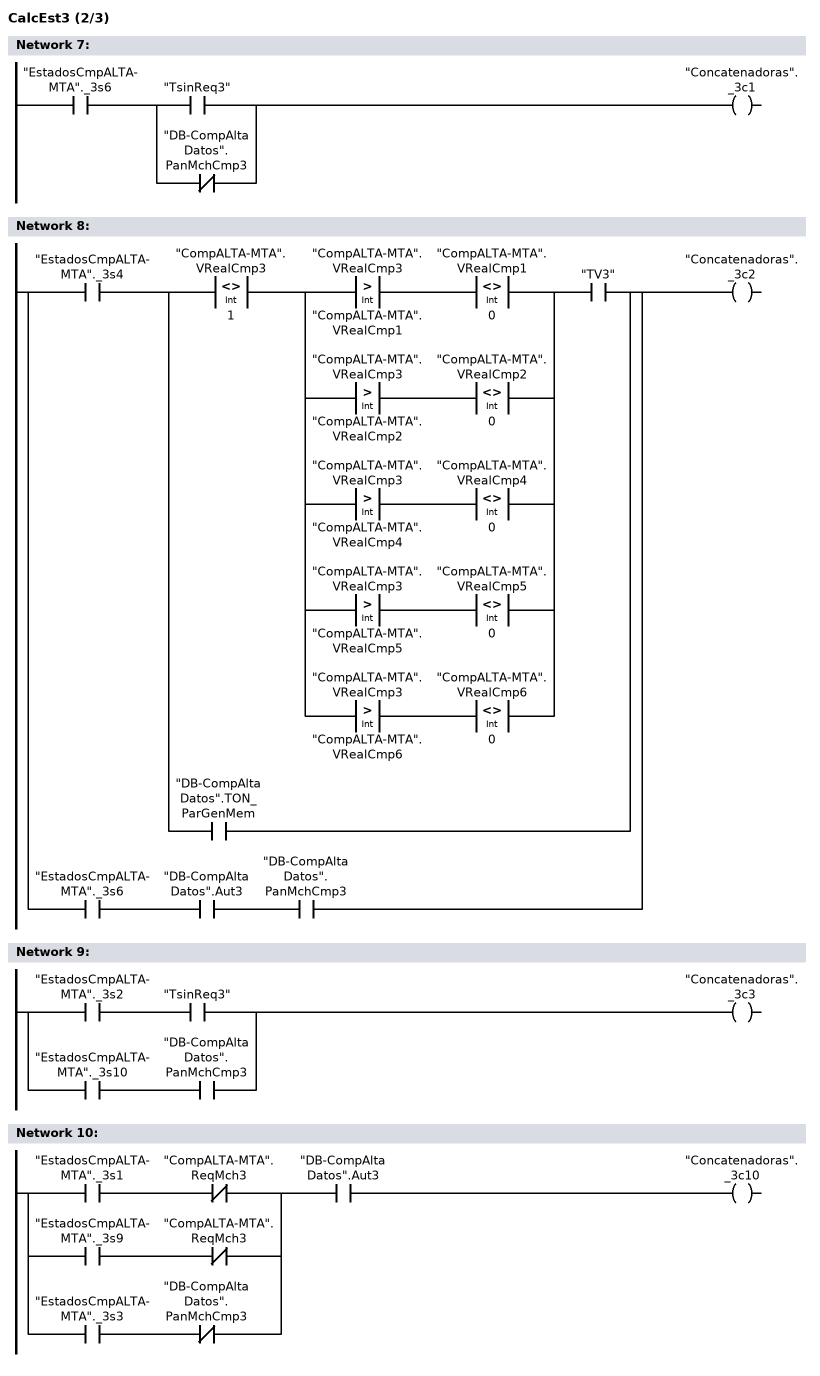
   RUNG wire#powerrail
      Contact( "EstadosCmpALTA-MTA"._3s6 )
      wire#w1
      Contact( "TsinReq3" )
      wire#w2
      Coil( "Concatenadoras"._3c1 )
   END_RUNG
   RUNG wire#w1
      I_Contact( "DB-CompAltaDatos".PanMchCmp3 )
   END_RUNG wire#w2
   // the same network as SCL:
   "Concatenadoras"._3c1 := "EstadosCmpALTA-MTA"._3s6 AND ("TsinReq3" OR NOT "DB-CompAltaDatos".PanMchCmp3);
END_REGION

REGION Network 8
   RUNG wire#powerrail
      Contact( "EstadosCmpALTA-MTA"._3s4 )
      wire#w1
      { S7_Templates := "SrcType := Int" } NE_Contact(in1 := "CompALTA-MTA".VRealCmp3, in2 := 1)
      wire#w2
      { S7_Templates := "SrcType := Int" } GT_Contact(in1 := "CompALTA-MTA".VRealCmp3, in2 := "CompALTA-MTA".VRealCmp1)
      { S7_Templates := "SrcType := Int" } NE_Contact(in1 := "CompALTA-MTA".VRealCmp1, in2 := 0)
      wire#w3
      Contact( "TV3" )
      wire#w4
      Coil( "Concatenadoras"._3c2 )
   END_RUNG
   RUNG wire#w2
      { S7_Templates := "SrcType := Int" } GT_Contact(in1 := "CompALTA-MTA".VRealCmp3, in2 := "CompALTA-MTA".VRealCmp2)
      { S7_Templates := "SrcType := Int" } NE_Contact(in1 := "CompALTA-MTA".VRealCmp2, in2 := 0)
   END_RUNG wire#w3
   RUNG wire#w2
      { S7_Templates := "SrcType := Int" } GT_Contact(in1 := "CompALTA-MTA".VRealCmp3, in2 := "CompALTA-MTA".VRealCmp4)
      { S7_Templates := "SrcType := Int" } NE_Contact(in1 := "CompALTA-MTA".VRealCmp4, in2 := 0)
   END_RUNG wire#w3
   RUNG wire#w2
      { S7_Templates := "SrcType := Int" } GT_Contact(in1 := "CompALTA-MTA".VRealCmp3, in2 := "CompALTA-MTA".VRealCmp5)
      { S7_Templates := "SrcType := Int" } NE_Contact(in1 := "CompALTA-MTA".VRealCmp5, in2 := 0)
   END_RUNG wire#w3
   RUNG wire#w2
      { S7_Templates := "SrcType := Int" } GT_Contact(in1 := "CompALTA-MTA".VRealCmp3, in2 := "CompALTA-MTA".VRealCmp6)
      { S7_Templates := "SrcType := Int" } NE_Contact(in1 := "CompALTA-MTA".VRealCmp6, in2 := 0)
   END_RUNG wire#w3
   RUNG wire#w1
      Contact( "DB-CompAltaDatos".TON_ParGenMem )
   END_RUNG wire#w4
   RUNG wire#powerrail
      Contact( "EstadosCmpALTA-MTA"._3s6 )
      Contact( "DB-CompAltaDatos".Aut3 )
      Contact( "DB-CompAltaDatos".PanMchCmp3 )
   END_RUNG wire#w4
   // the same network as SCL:
   "Concatenadoras"._3c2 := ("EstadosCmpALTA-MTA"._3s4 AND ((("CompALTA-MTA".VRealCmp3 <> 1) AND ((("CompALTA-MTA".VRealCmp3 > "CompALTA-MTA".VRealCmp1) AND ("CompALTA-MTA".VRealCmp1 <> 0)) OR (("CompALTA-MTA".VRealCmp3 > "CompALTA-MTA".VRealCmp2) AND ("CompALTA-MTA".VRealCmp2 <> 0)) OR (("CompALTA-MTA".VRealCmp3 > "CompALTA-MTA".VRealCmp4) AND ("CompALTA-MTA".VRealCmp4 <> 0)) OR (("CompALTA-MTA".VRealCmp3 > "CompALTA-MTA".VRealCmp5) AND ("CompALTA-MTA".VRealCmp5 <> 0)) OR (("CompALTA-MTA".VRealCmp3 > "CompALTA-MTA".VRealCmp6) AND ("CompALTA-MTA".VRealCmp6 <> 0))) AND "TV3") OR "DB-CompAltaDatos".TON_ParGenMem)) OR ("EstadosCmpALTA-MTA"._3s6 AND "DB-CompAltaDatos".Aut3 AND "DB-CompAltaDatos".PanMchCmp3);
END_REGION

REGION Network 9
   RUNG wire#powerrail
      Contact( "EstadosCmpALTA-MTA"._3s2 )
      Contact( "TsinReq3" )
      wire#w1
      Coil( "Concatenadoras"._3c3 )
   END_RUNG
   RUNG wire#powerrail
      Contact( "EstadosCmpALTA-MTA"._3s10 )
      Contact( "DB-CompAltaDatos".PanMchCmp3 )
   END_RUNG wire#w1
   // the same network as SCL:
   "Concatenadoras"._3c3 := ("EstadosCmpALTA-MTA"._3s2 AND "TsinReq3") OR ("EstadosCmpALTA-MTA"._3s10 AND "DB-CompAltaDatos".PanMchCmp3);
END_REGION

REGION Network 10
   RUNG wire#powerrail
      Contact( "EstadosCmpALTA-MTA"._3s1 )
      I_Contact( "CompALTA-MTA".ReqMch3 )
      wire#w1
      Contact( "DB-CompAltaDatos".Aut3 )
      Coil( "Concatenadoras"._3c10 )
   END_RUNG
   RUNG wire#powerrail
      Contact( "EstadosCmpALTA-MTA"._3s9 )
      I_Contact( "CompALTA-MTA".ReqMch3 )
   END_RUNG wire#w1
   RUNG wire#powerrail
      Contact( "EstadosCmpALTA-MTA"._3s3 )
      I_Contact( "DB-CompAltaDatos".PanMchCmp3 )
   END_RUNG wire#w1
   // the same network as SCL:
   "Concatenadoras"._3c10 := (("EstadosCmpALTA-MTA"._3s1 AND NOT "CompALTA-MTA".ReqMch3) OR ("EstadosCmpALTA-MTA"._3s9 AND NOT "CompALTA-MTA".ReqMch3) OR ("EstadosCmpALTA-MTA"._3s3 AND NOT "DB-CompAltaDatos".PanMchCmp3)) AND "DB-CompAltaDatos".Aut3;
END_REGION

REGION Network 11
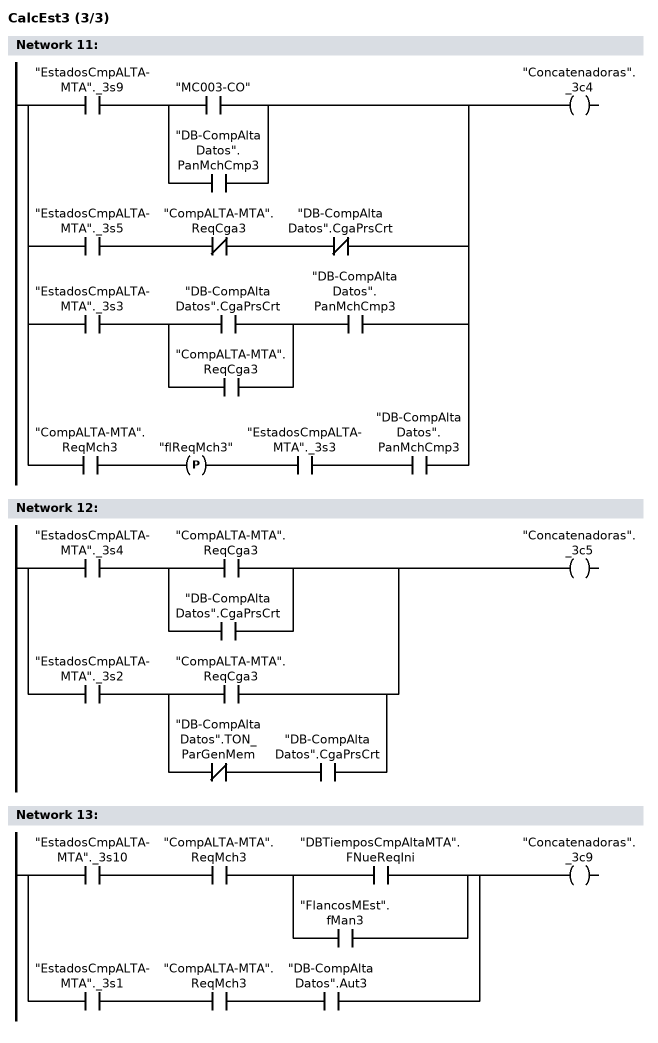
   RUNG wire#powerrail
      Contact( "EstadosCmpALTA-MTA"._3s9 )
      wire#w1
      Contact( "MC003-CO" )
      wire#w2
      Coil( "Concatenadoras"._3c4 )
   END_RUNG
   RUNG wire#w1
      Contact( "DB-CompAltaDatos".PanMchCmp3 )
   END_RUNG wire#w2
   RUNG wire#powerrail
      Contact( "EstadosCmpALTA-MTA"._3s5 )
      I_Contact( "CompALTA-MTA".ReqCga3 )
      I_Contact( "DB-CompAltaDatos".CgaPrsCrt )
   END_RUNG wire#w2
   RUNG wire#powerrail
      Contact( "EstadosCmpALTA-MTA"._3s3 )
      wire#w3
      Contact( "DB-CompAltaDatos".CgaPrsCrt )
      wire#w4
      Contact( "DB-CompAltaDatos".PanMchCmp3 )
   END_RUNG wire#w2
   RUNG wire#w3
      Contact( "CompALTA-MTA".ReqCga3 )
   END_RUNG wire#w4
   RUNG wire#powerrail
      Contact( "CompALTA-MTA".ReqMch3 )
      P_Trig( "flReqMch3" )
      Contact( "EstadosCmpALTA-MTA"._3s3 )
      Contact( "DB-CompAltaDatos".PanMchCmp3 )
   END_RUNG wire#w2
   // the same network as SCL:
   #_w1 := "CompALTA-MTA".ReqMch3 AND NOT "flReqMch3";   // rising edge
   "flReqMch3" := "CompALTA-MTA".ReqMch3;
   "Concatenadoras"._3c4 := ("EstadosCmpALTA-MTA"._3s9 AND ("MC003-CO" OR "DB-CompAltaDatos".PanMchCmp3)) OR ("EstadosCmpALTA-MTA"._3s5 AND NOT "CompALTA-MTA".ReqCga3 AND NOT "DB-CompAltaDatos".CgaPrsCrt) OR ("EstadosCmpALTA-MTA"._3s3 AND ("DB-CompAltaDatos".CgaPrsCrt OR "CompALTA-MTA".ReqCga3) AND "DB-CompAltaDatos".PanMchCmp3) OR (#_w1 AND "EstadosCmpALTA-MTA"._3s3 AND "DB-CompAltaDatos".PanMchCmp3);
END_REGION

REGION Network 12
   RUNG wire#powerrail
      Contact( "EstadosCmpALTA-MTA"._3s4 )
      wire#w1
      Contact( "CompALTA-MTA".ReqCga3 )
      wire#w2
      Coil( "Concatenadoras"._3c5 )
   END_RUNG
   RUNG wire#w1
      Contact( "DB-CompAltaDatos".CgaPrsCrt )
   END_RUNG wire#w2
   RUNG wire#powerrail
      Contact( "EstadosCmpALTA-MTA"._3s2 )
      wire#w3
      Contact( "CompALTA-MTA".ReqCga3 )
   END_RUNG wire#w2
   RUNG wire#w3
      I_Contact( "DB-CompAltaDatos".TON_ParGenMem )
      Contact( "DB-CompAltaDatos".CgaPrsCrt )
   END_RUNG wire#w2
   // the same network as SCL:
   "Concatenadoras"._3c5 := ("EstadosCmpALTA-MTA"._3s4 AND ("CompALTA-MTA".ReqCga3 OR "DB-CompAltaDatos".CgaPrsCrt)) OR ("EstadosCmpALTA-MTA"._3s2 AND ("CompALTA-MTA".ReqCga3 OR (NOT "DB-CompAltaDatos".TON_ParGenMem AND "DB-CompAltaDatos".CgaPrsCrt)));
END_REGION

REGION Network 13
   RUNG wire#powerrail
      Contact( "EstadosCmpALTA-MTA"._3s10 )
      Contact( "CompALTA-MTA".ReqMch3 )
      wire#w1
      Contact( "DBTiemposCmpAltaMTA".FNueReqIni )
      wire#w2
      Coil( "Concatenadoras"._3c9 )
   END_RUNG
   RUNG wire#w1
      Contact( "FlancosMEst".fMan3 )
   END_RUNG wire#w2
   RUNG wire#powerrail
      Contact( "EstadosCmpALTA-MTA"._3s1 )
      Contact( "CompALTA-MTA".ReqMch3 )
      Contact( "DB-CompAltaDatos".Aut3 )
   END_RUNG wire#w2
   // the same network as SCL:
   "Concatenadoras"._3c9 := ("EstadosCmpALTA-MTA"._3s10 AND "CompALTA-MTA".ReqMch3 AND ("DBTiemposCmpAltaMTA".FNueReqIni OR "FlancosMEst".fMan3)) OR ("EstadosCmpALTA-MTA"._3s1 AND "CompALTA-MTA".ReqMch3 AND "DB-CompAltaDatos".Aut3);
END_REGION

REGION Network 14 (STL)
         CALL  "FC_MAQ_EST_16"
         ( IN0  := %DB127.DBW4,
           IN1  := %DB128.DBW4,
           OUT2 := "ErrPMQ3",
           OUT3 := "ErrCMQ3",
           IO4  := %DB120.DBW4
         );
         NOP   0;
END_REGION

REGION Network 15 (STL)
         CALL  "FC-ANIM-CMP"
         ( IN0  := %DB120.DBW4,
           OUT1 := "CompALTA-MTA".AnimCMP3
         );
         NOP   0;
END_REGION
END_FUNCTION

FUNCTION "CalcEst4" : Void   // FC39, LAD
{ S7_Optimized_Access := 'FALSE' }
VERSION : 0.1
   VAR_TEMP   // added for the SCL form of the ladder/FBD networks
      _w1 : Bool;
   END_VAR
BEGIN

REGION Network 1
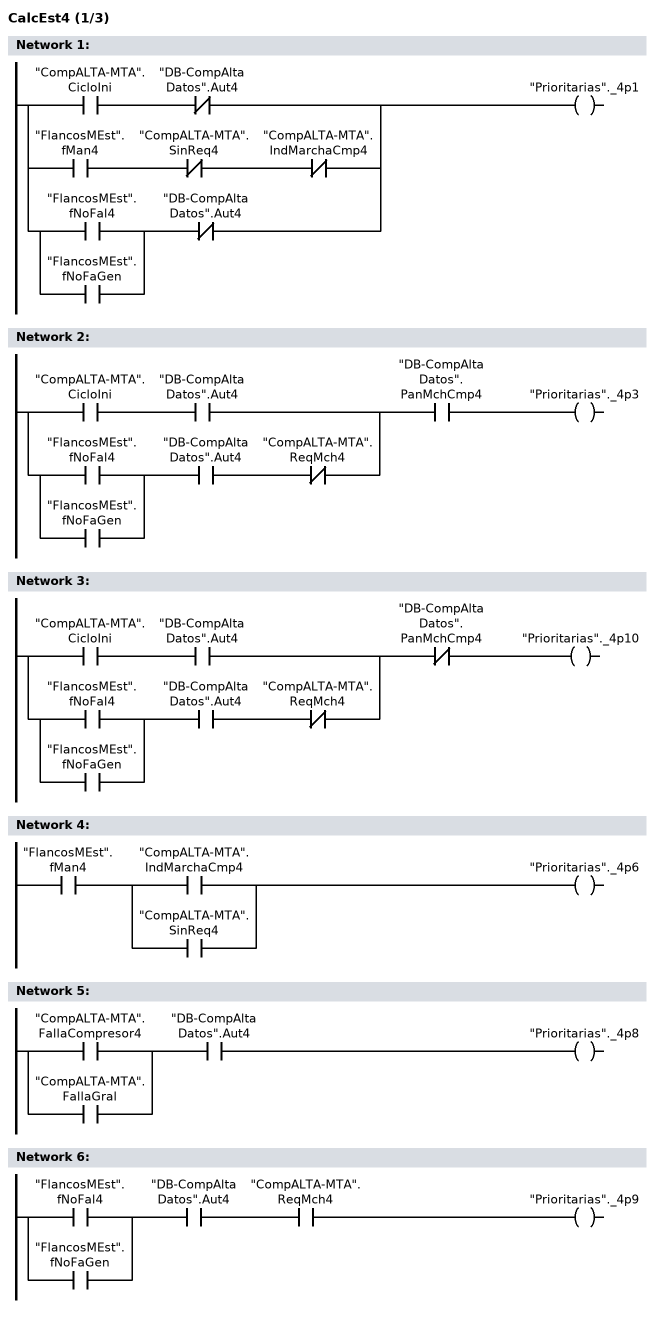
   RUNG wire#powerrail
      Contact( "CompALTA-MTA".CicloIni )
      I_Contact( "DB-CompAltaDatos".Aut4 )
      wire#w1
      Coil( "Prioritarias"._4p1 )
   END_RUNG
   RUNG wire#powerrail
      Contact( "FlancosMEst".fMan4 )
      I_Contact( "CompALTA-MTA".SinReq4 )
      I_Contact( "CompALTA-MTA".IndMarchaCmp4 )
   END_RUNG wire#w1
   RUNG wire#powerrail
      Contact( "FlancosMEst".fNoFal4 )
      wire#w2
      I_Contact( "DB-CompAltaDatos".Aut4 )
   END_RUNG wire#w1
   RUNG wire#powerrail
      Contact( "FlancosMEst".fNoFaGen )
   END_RUNG wire#w2
   // the same network as SCL:
   "Prioritarias"._4p1 := ("CompALTA-MTA".CicloIni AND NOT "DB-CompAltaDatos".Aut4) OR ("FlancosMEst".fMan4 AND NOT "CompALTA-MTA".SinReq4 AND NOT "CompALTA-MTA".IndMarchaCmp4) OR (("FlancosMEst".fNoFal4 OR "FlancosMEst".fNoFaGen) AND NOT "DB-CompAltaDatos".Aut4);
END_REGION

REGION Network 2
   RUNG wire#powerrail
      Contact( "CompALTA-MTA".CicloIni )
      Contact( "DB-CompAltaDatos".Aut4 )
      wire#w1
      Contact( "DB-CompAltaDatos".PanMchCmp4 )
      Coil( "Prioritarias"._4p3 )
   END_RUNG
   RUNG wire#powerrail
      Contact( "FlancosMEst".fNoFal4 )
      wire#w2
      Contact( "DB-CompAltaDatos".Aut4 )
      I_Contact( "CompALTA-MTA".ReqMch4 )
   END_RUNG wire#w1
   RUNG wire#powerrail
      Contact( "FlancosMEst".fNoFaGen )
   END_RUNG wire#w2
   // the same network as SCL:
   "Prioritarias"._4p3 := (("CompALTA-MTA".CicloIni AND "DB-CompAltaDatos".Aut4) OR (("FlancosMEst".fNoFal4 OR "FlancosMEst".fNoFaGen) AND "DB-CompAltaDatos".Aut4 AND NOT "CompALTA-MTA".ReqMch4)) AND "DB-CompAltaDatos".PanMchCmp4;
END_REGION

REGION Network 3
   RUNG wire#powerrail
      Contact( "CompALTA-MTA".CicloIni )
      Contact( "DB-CompAltaDatos".Aut4 )
      wire#w1
      I_Contact( "DB-CompAltaDatos".PanMchCmp4 )
      Coil( "Prioritarias"._4p10 )
   END_RUNG
   RUNG wire#powerrail
      Contact( "FlancosMEst".fNoFal4 )
      wire#w2
      Contact( "DB-CompAltaDatos".Aut4 )
      I_Contact( "CompALTA-MTA".ReqMch4 )
   END_RUNG wire#w1
   RUNG wire#powerrail
      Contact( "FlancosMEst".fNoFaGen )
   END_RUNG wire#w2
   // the same network as SCL:
   "Prioritarias"._4p10 := (("CompALTA-MTA".CicloIni AND "DB-CompAltaDatos".Aut4) OR (("FlancosMEst".fNoFal4 OR "FlancosMEst".fNoFaGen) AND "DB-CompAltaDatos".Aut4 AND NOT "CompALTA-MTA".ReqMch4)) AND NOT "DB-CompAltaDatos".PanMchCmp4;
END_REGION

REGION Network 4
   RUNG wire#powerrail
      Contact( "FlancosMEst".fMan4 )
      wire#w1
      Contact( "CompALTA-MTA".IndMarchaCmp4 )
      wire#w2
      Coil( "Prioritarias"._4p6 )
   END_RUNG
   RUNG wire#w1
      Contact( "CompALTA-MTA".SinReq4 )
   END_RUNG wire#w2
   // the same network as SCL:
   "Prioritarias"._4p6 := "FlancosMEst".fMan4 AND ("CompALTA-MTA".IndMarchaCmp4 OR "CompALTA-MTA".SinReq4);
END_REGION

REGION Network 5
   RUNG wire#powerrail
      Contact( "CompALTA-MTA".FallaCompresor4 )
      wire#w1
      Contact( "DB-CompAltaDatos".Aut4 )
      Coil( "Prioritarias"._4p8 )
   END_RUNG
   RUNG wire#powerrail
      Contact( "CompALTA-MTA".FallaGral )
   END_RUNG wire#w1
   // the same network as SCL:
   "Prioritarias"._4p8 := ("CompALTA-MTA".FallaCompresor4 OR "CompALTA-MTA".FallaGral) AND "DB-CompAltaDatos".Aut4;
END_REGION

REGION Network 6
   RUNG wire#powerrail
      Contact( "FlancosMEst".fNoFal4 )
      wire#w1
      Contact( "DB-CompAltaDatos".Aut4 )
      Contact( "CompALTA-MTA".ReqMch4 )
      Coil( "Prioritarias"._4p9 )
   END_RUNG
   RUNG wire#powerrail
      Contact( "FlancosMEst".fNoFaGen )
   END_RUNG wire#w1
   // the same network as SCL:
   "Prioritarias"._4p9 := ("FlancosMEst".fNoFal4 OR "FlancosMEst".fNoFaGen) AND "DB-CompAltaDatos".Aut4 AND "CompALTA-MTA".ReqMch4;
END_REGION

REGION Network 7
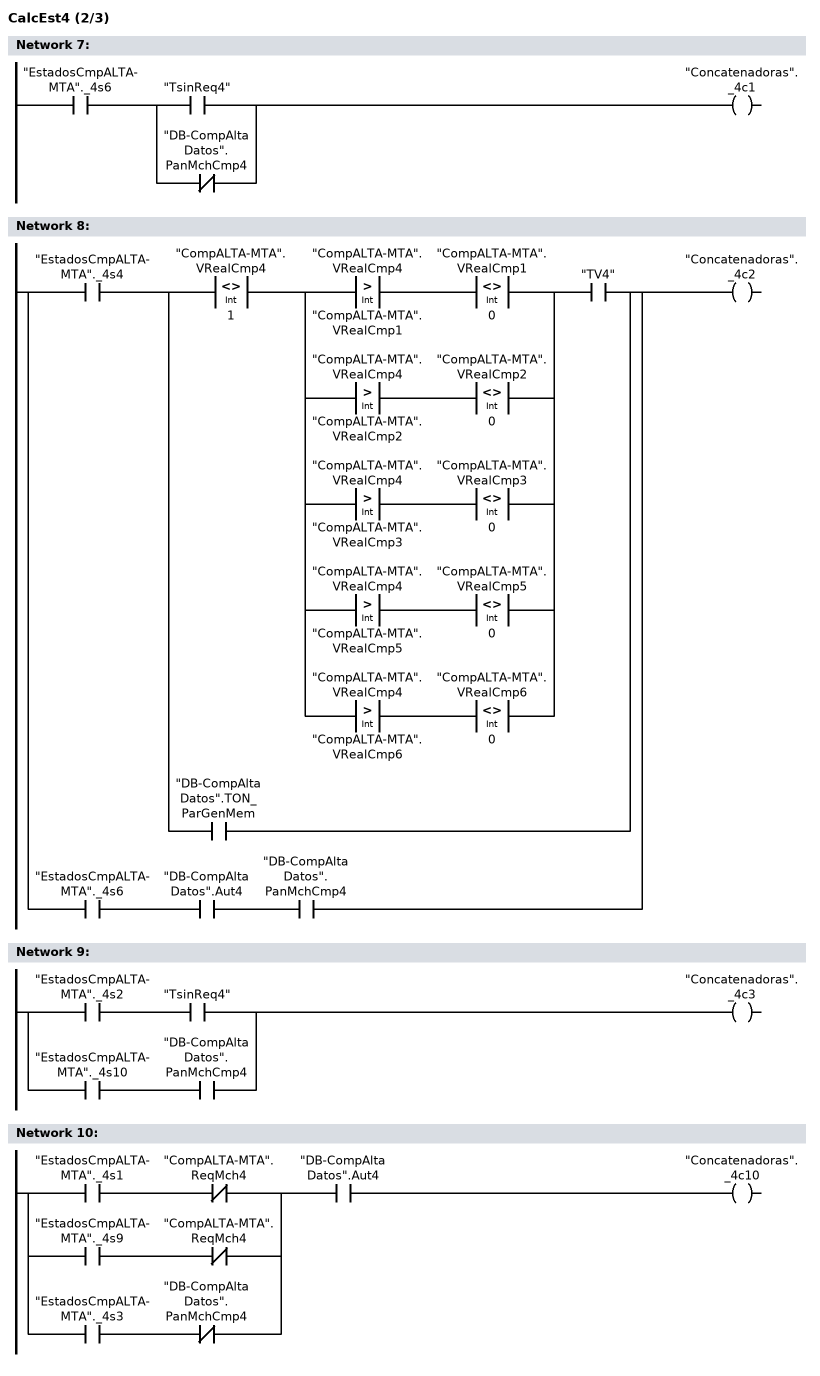
   RUNG wire#powerrail
      Contact( "EstadosCmpALTA-MTA"._4s6 )
      wire#w1
      Contact( "TsinReq4" )
      wire#w2
      Coil( "Concatenadoras"._4c1 )
   END_RUNG
   RUNG wire#w1
      I_Contact( "DB-CompAltaDatos".PanMchCmp4 )
   END_RUNG wire#w2
   // the same network as SCL:
   "Concatenadoras"._4c1 := "EstadosCmpALTA-MTA"._4s6 AND ("TsinReq4" OR NOT "DB-CompAltaDatos".PanMchCmp4);
END_REGION

REGION Network 8
   RUNG wire#powerrail
      Contact( "EstadosCmpALTA-MTA"._4s4 )
      wire#w1
      { S7_Templates := "SrcType := Int" } NE_Contact(in1 := "CompALTA-MTA".VRealCmp4, in2 := 1)
      wire#w2
      { S7_Templates := "SrcType := Int" } GT_Contact(in1 := "CompALTA-MTA".VRealCmp4, in2 := "CompALTA-MTA".VRealCmp1)
      { S7_Templates := "SrcType := Int" } NE_Contact(in1 := "CompALTA-MTA".VRealCmp1, in2 := 0)
      wire#w3
      Contact( "TV4" )
      wire#w4
      Coil( "Concatenadoras"._4c2 )
   END_RUNG
   RUNG wire#w2
      { S7_Templates := "SrcType := Int" } GT_Contact(in1 := "CompALTA-MTA".VRealCmp4, in2 := "CompALTA-MTA".VRealCmp2)
      { S7_Templates := "SrcType := Int" } NE_Contact(in1 := "CompALTA-MTA".VRealCmp2, in2 := 0)
   END_RUNG wire#w3
   RUNG wire#w2
      { S7_Templates := "SrcType := Int" } GT_Contact(in1 := "CompALTA-MTA".VRealCmp4, in2 := "CompALTA-MTA".VRealCmp3)
      { S7_Templates := "SrcType := Int" } NE_Contact(in1 := "CompALTA-MTA".VRealCmp3, in2 := 0)
   END_RUNG wire#w3
   RUNG wire#w2
      { S7_Templates := "SrcType := Int" } GT_Contact(in1 := "CompALTA-MTA".VRealCmp4, in2 := "CompALTA-MTA".VRealCmp5)
      { S7_Templates := "SrcType := Int" } NE_Contact(in1 := "CompALTA-MTA".VRealCmp5, in2 := 0)
   END_RUNG wire#w3
   RUNG wire#w2
      { S7_Templates := "SrcType := Int" } GT_Contact(in1 := "CompALTA-MTA".VRealCmp4, in2 := "CompALTA-MTA".VRealCmp6)
      { S7_Templates := "SrcType := Int" } NE_Contact(in1 := "CompALTA-MTA".VRealCmp6, in2 := 0)
   END_RUNG wire#w3
   RUNG wire#w1
      Contact( "DB-CompAltaDatos".TON_ParGenMem )
   END_RUNG wire#w4
   RUNG wire#powerrail
      Contact( "EstadosCmpALTA-MTA"._4s6 )
      Contact( "DB-CompAltaDatos".Aut4 )
      Contact( "DB-CompAltaDatos".PanMchCmp4 )
   END_RUNG wire#w4
   // the same network as SCL:
   "Concatenadoras"._4c2 := ("EstadosCmpALTA-MTA"._4s4 AND ((("CompALTA-MTA".VRealCmp4 <> 1) AND ((("CompALTA-MTA".VRealCmp4 > "CompALTA-MTA".VRealCmp1) AND ("CompALTA-MTA".VRealCmp1 <> 0)) OR (("CompALTA-MTA".VRealCmp4 > "CompALTA-MTA".VRealCmp2) AND ("CompALTA-MTA".VRealCmp2 <> 0)) OR (("CompALTA-MTA".VRealCmp4 > "CompALTA-MTA".VRealCmp3) AND ("CompALTA-MTA".VRealCmp3 <> 0)) OR (("CompALTA-MTA".VRealCmp4 > "CompALTA-MTA".VRealCmp5) AND ("CompALTA-MTA".VRealCmp5 <> 0)) OR (("CompALTA-MTA".VRealCmp4 > "CompALTA-MTA".VRealCmp6) AND ("CompALTA-MTA".VRealCmp6 <> 0))) AND "TV4") OR "DB-CompAltaDatos".TON_ParGenMem)) OR ("EstadosCmpALTA-MTA"._4s6 AND "DB-CompAltaDatos".Aut4 AND "DB-CompAltaDatos".PanMchCmp4);
END_REGION

REGION Network 9
   RUNG wire#powerrail
      Contact( "EstadosCmpALTA-MTA"._4s2 )
      Contact( "TsinReq4" )
      wire#w1
      Coil( "Concatenadoras"._4c3 )
   END_RUNG
   RUNG wire#powerrail
      Contact( "EstadosCmpALTA-MTA"._4s10 )
      Contact( "DB-CompAltaDatos".PanMchCmp4 )
   END_RUNG wire#w1
   // the same network as SCL:
   "Concatenadoras"._4c3 := ("EstadosCmpALTA-MTA"._4s2 AND "TsinReq4") OR ("EstadosCmpALTA-MTA"._4s10 AND "DB-CompAltaDatos".PanMchCmp4);
END_REGION
